
                 // ---------------------------------------------------
                 // GLOBAL
                 // If not local variable then check if global
                 // ---------------------------------------------------
                 // Variable definition should look like this:
                 // DEF GLOBAL DINT myVar_1 --> Create global integer var "myVar_1" 
                 //
                 // Token:
                 // [1] myVar_1
                 // [2]
                 // [3] DINT
                 // [4]
                 // [5] GLOBAL
                 // [6] 
                 // [7] DEF

                 // Init temp
                 #tempGlobal := FALSE;

                 // Check if number of token fits
                 IF #statTokenizedLine.numberOfToken = #statGlobalVariableDefinition.tokenizedString.numberOfToken THEN
                   // Set state initially --> Is overwritten in for loop
                   #statStateIntern := #STATE_LINE_IS_VAR_DEF;
                   #tempGlobal := TRUE;

                   // Check token of line to fit var declaration
                   FOR #tempCounter := 1 TO #statTokenizedLine.numberOfToken DO
                     // Skip name and type token
                     IF #tempCounter = #statGlobalVariableDefinition.nameTokenNumber
                       OR #tempCounter = #statGlobalVariableDefinition.typeTokenNumber
                     THEN
                       CONTINUE;
                       // Check the other keywords
                     ELSIF #statTokenizedLine.lineToken[#tempCounter] <> #statGlobalVariableDefinition.tokenizedString.lineToken[#tempCounter] THEN
                       // Mismatch between defintion and line 
                       // --> Not a variable definition
                       #statStateIntern := #STATE_IS_LINE_LABEL;
                       #tempGlobal := FALSE;
                       EXIT;
                     END_IF;
                   END_FOR;
                 ELSE
                   // Number of token does not fit
                   // Parse normal line
                   // Next step 
                   #statStateIntern := #STATE_IS_LINE_LABEL;
                   #tempGlobal := FALSE;
                 END_IF;

                 // Only check for local if not global
                 IF #tempGlobal = FALSE THEN
                   // ---------------------------------------------------
                   // LOCAL
                   // ---------------------------------------------------
                   // Variable definition should look like this:
                   // DEF DINT myVar_1 --> Create local integer var "myVar_1" 
                   //
                   // Token:
                   // [1] myVar_1
                   // [2]
                   // [3] DINT
                   // [4]
                   // [5] DEF

                   // Check if number of token fits
                   IF #statTokenizedLine.numberOfToken = #statLocalVariableDefinition.tokenizedString.numberOfToken THEN
                     // Set state initially --> Is overwritten in for loop
                     #statStateIntern := #STATE_LINE_IS_VAR_DEF;

                     // Check token of line to fit var declaration
                     FOR #tempCounter := 1 TO #statTokenizedLine.numberOfToken DO
                       // Skip name and type token
                       IF #tempCounter = #statLocalVariableDefinition.nameTokenNumber
                         OR #tempCounter = #statLocalVariableDefinition.typeTokenNumber
                       THEN
                         CONTINUE;
                         // Check the other keywords
                       ELSIF #statTokenizedLine.lineToken[#tempCounter] <> #statLocalVariableDefinition.tokenizedString.lineToken[#tempCounter] THEN
                         // Mismatch between defintion and line 
                         // --> Not a variable definition
                         #statStateIntern := #STATE_IS_LINE_LABEL;
                         EXIT;
                       END_IF;
                     END_FOR;
                   ELSE
                     // Number of token does not fit
                     // Parse normal line
                     // Next step 
                     #statStateIntern := #STATE_IS_LINE_LABEL;
                   END_IF;
                 END_IF;

               END_IF;

             END_REGION IS_LINE_VARIABLE_DEFINITION


             // ------------------------------------------------------------------------------------------
             // Line is variable definition
             // Line contains a variable definition like "DEF DINT myVar_1"
             // Go to STATE_LINE_PARSED
             // ------------------------------------------------------------------------------------------ 
             REGION LINE_IS_VARIABLE_DEFINITION
               IF #statStateIntern = #STATE_LINE_IS_VAR_DEF
               THEN
                 // Variable definition should look like this:
                 // DEF DINT myVar_1 --> Create local integer var "myVar_1" 
                 // Token:
                 // [1] myVar_1
                 // [2]
                 // [3] DINT
                 // [4]
                 // [5] DEF

                 // Check name to not be a number only!
                 IF NOT "LKinLang_IsTokenNumberInclSign"(#statTokenizedLine.lineToken[#statLocalVariableDefinition.nameTokenNumber]) THEN

                   // Check if name already exists as LABEL!
                   FOR #tempVarIndex := 1 TO #statLabelList.numberOfLabels DO
                     IF #statLabelList.labels[#tempVarIndex].labelName = #statTokenizedLine.lineToken[#statLocalVariableDefinition.nameTokenNumber] THEN
                       // Error: Variable already exists as label
                       #statStatus := #ERR_PARSING;
                       #statStateIntern := #STATE_ERROR;
                       #statErrorString := CONCAT(IN1 := #statErrorString, IN2 := 'Error: Variable already exists as label');
                       #statErrorString := CONCAT(IN1 := #statErrorString, IN2 := '; Line: ');
                       #statErrorString := CONCAT(IN1 := #statErrorString, IN2 := UDINT_TO_STRING(#statTokenizedLine.lineNo));
                       EXIT;
                     END_IF;
                   END_FOR;

                   // Check if name is a keyword
                   IF "LKinLang_IsTokenKeyWord"(token := #statTokenizedLine.lineToken[#statLocalVariableDefinition.nameTokenNumber], keyToken := #statKeyToken) THEN
                     // Error: Variable name can not be a keyword
                     #statStatus := #ERR_PARSING;
                     #statStateIntern := #STATE_ERROR;
                     #statErrorString := CONCAT(IN1 := #statErrorString, IN2 := 'Error: Variable name must not be a keyword');
                     #statErrorString := CONCAT(IN1 := #statErrorString, IN2 := '; Line: ');
                     #statErrorString := CONCAT(IN1 := #statErrorString, IN2 := UDINT_TO_STRING(#statTokenizedLine.lineNo));
                     EXIT;
                   END_IF;

                   // Check if name is a parameter 
                   FOR #tempVarIndex := 1 TO "LKINLANG_MAX_NUMBER_OF_PARAMETERS" DO
                     IF #statParameterLookUpTable[#tempVarIndex].parameterNameString = #statTokenizedLine.lineToken[#statLocalVariableDefinition.nameTokenNumber] THEN
                       // Error: Variable name can not be a keyword
                       #statStatus := #ERR_PARSING;
                       #statStateIntern := #STATE_ERROR;
                       #statErrorString := CONCAT(IN1 := #statErrorString, IN2 := 'Error: Variable name must not be a keyword');
                       #statErrorString := CONCAT(IN1 := #statErrorString, IN2 := '; Line: ');
                       #statErrorString := CONCAT(IN1 := #statErrorString, IN2 := UDINT_TO_STRING(#statTokenizedLine.lineNo));
                       EXIT;
                     END_IF;
                   END_FOR;

                   // Check if error occurred before
                   IF #statStateIntern <> #STATE_ERROR THEN
                     // Create local variable
                     // Imcrement local var counter
                     #statVarRefList.numberOfReferences += 1;

                     IF #statVarRefList.numberOfReferences > "LKINLANG_NUMBER_OF_VAR_REFS" THEN
                       // Error: Max number of variable references reached
                       #statStatus := #ERR_PARSING;
                       #statStateIntern := #STATE_ERROR;
                       #statErrorString := CONCAT(IN1 := #statErrorString, IN2 := 'Error: Overflow VarRefList; Increase NUMBER_OF_VAR_REFS');
                       #statErrorString := CONCAT(IN1 := #statErrorString, IN2 := '; Line: ');
                       #statErrorString := CONCAT(IN1 := #statErrorString, IN2 := UDINT_TO_STRING(#statTokenizedLine.lineNo));
                       EXIT;
                     ELSE
                       // Set step here because changing to error state could happen afterwards
                       // Next step --> Line finished
                       #statStateIntern := #STATE_LINE_PARSED;

                       // Copy name to table
                       #statVarRefList.references[#statVarRefList.numberOfReferences].name := #statTokenizedLine.lineToken[#statLocalVariableDefinition.nameTokenNumber];

                       // Check and set scope 
                       // Preset the scope to main
                       IF #tempGlobal = TRUE THEN
                         #statVarRefList.references[#statVarRefList.numberOfReferences].scope := 2; // Global var in main prg
                       ELSE
                         #statVarRefList.references[#statVarRefList.numberOfReferences].scope := 1; // Local var in main prg
                       END_IF;

                       // Iterate over subProgramList and check where we are currently
                       FOR #tempCounter := 1 TO #statSubPrgList.numberOfSubPrgs DO
                         IF #statTokenizedLine.lineNo > #statSubPrgList.subPrgs[#tempCounter].lineNumberStart
                           AND #statTokenizedLine.lineNo < #statSubPrgList.subPrgs[#tempCounter].lineNumberEnd
                         THEN
                           #statVarRefList.references[#statVarRefList.numberOfReferences].scope := #tempCounter * 10; // Local var in sub prg 
                           EXIT;
                         ELSIF #statTokenizedLine.lineNo < #statSubPrgList.subPrgs[#tempCounter].lineNumberStart THEN // Check if the current line number is smaller than the start of a sub --> Exit earlier
                           EXIT;
                         ELSE
                           CONTINUE;
                         END_IF;
                       END_FOR;

                       // Check if Global is allowed 
                       IF #tempGlobal = TRUE
                         AND #statVarRefList.references[#statVarRefList.numberOfReferences].scope >= 10
                       THEN
                         // Error: Not allowed to declare global in sub
                         #statStatus := #ERR_PARSING;
                         #statStateIntern := #STATE_ERROR;
                         #statErrorString := CONCAT(IN1 := #statErrorString, IN2 := 'Error: Declaring global variable in subprogram not allowed');
                         #statErrorString := CONCAT(IN1 := #statErrorString, IN2 := '; Line: ');
                         #statErrorString := CONCAT(IN1 := #statErrorString, IN2 := UDINT_TO_STRING(#statTokenizedLine.lineNo));
                         EXIT;
                       END_IF;

                       // Check if name already exists!
                       FOR #tempVarIndex := 1 TO #statVarRefList.numberOfReferences - 1 DO // exclude current entry
                         IF #statVarRefList.references[#tempVarIndex].name = #statVarRefList.references[#statVarRefList.numberOfReferences].name
                           AND #statVarRefList.references[#tempVarIndex].scope = #statVarRefList.references[#statVarRefList.numberOfReferences].scope
                         THEN
                           // Error: Variable already exists
                           #statStatus := #ERR_PARSING;
                           #statStateIntern := #STATE_ERROR;
                           #statErrorString := CONCAT(IN1 := #statErrorString, IN2 := 'Error: Variable already exists');
                           #statErrorString := CONCAT(IN1 := #statErrorString, IN2 := '; Line: ');
                           #statErrorString := CONCAT(IN1 := #statErrorString, IN2 := UDINT_TO_STRING(#statTokenizedLine.lineNo));
                           EXIT;
                         END_IF;
                       END_FOR;

                       // Decide type of variable
                       IF #statTokenizedLine.lineToken[#statLocalVariableDefinition.typeTokenNumber] = #statKeyToken.tokenBool THEN
                         #statVarRefList.references[#statVarRefList.numberOfReferences].type := "LKINLANG_VAR_TYPE_LOCAL_BOOL";
                         #statVariables.boolCounter += 1;
                         IF #statVariables.boolCounter > "LKINLANG_NUMBER_OF_LOCAL_BOOL" THEN
                           // Error too many local boolean
                           #statStatus := #ERR_PARSING;
                           #statStateIntern := #STATE_ERROR;
                           #statErrorString := CONCAT(IN1 := #statErrorString, IN2 := 'Error: Overflow local Bool; Increase "LKINLANG_NUMBER_OF_LOCAL_BOOL"');
                           #statErrorString := CONCAT(IN1 := #statErrorString, IN2 := '; Line: ');
                           #statErrorString := CONCAT(IN1 := #statErrorString, IN2 := UDINT_TO_STRING(#statTokenizedLine.lineNo));
                           EXIT;
                         ELSE
                           #statVarRefList.references[#statVarRefList.numberOfReferences].index := #statVariables.boolCounter;
                           #statVariables.boolean[#statVariables.boolCounter] := FALSE;
                         END_IF;
                       ELSIF #statTokenizedLine.lineToken[#statLocalVariableDefinition.typeTokenNumber] = #statKeyToken.tokenDInt THEN
                         #statVarRefList.references[#statVarRefList.numberOfReferences].type := "LKINLANG_VAR_TYPE_LOCAL_DINT";
                         #statVariables.dintCounter += 1;
                         IF #statVariables.dintCounter > "LKINLANG_NUMBER_OF_LOCAL_DINT" THEN
                           // Error too many local DInt
                           #statStatus := #ERR_PARSING;
                           #statStateIntern := #STATE_ERROR;
                           #statErrorString := CONCAT(IN1 := #statErrorString, IN2 := 'Error: Overflow local DInt; Increase "LKINLANG_NUMBER_OF_LOCAL_DINT"');
                           #statErrorString := CONCAT(IN1 := #statErrorString, IN2 := '; Line: ');
                           #statErrorString := CONCAT(IN1 := #statErrorString, IN2 := UDINT_TO_STRING(#statTokenizedLine.lineNo));
                           EXIT;
                         ELSE
                           #statVarRefList.references[#statVarRefList.numberOfReferences].index := #statVariables.dintCounter;
                           #statVariables.dints[#statVariables.dintCounter] := 0;
                         END_IF;
                       ELSIF #statTokenizedLine.lineToken[#statLocalVariableDefinition.typeTokenNumber] = #statKeyToken.tokenLReal THEN
                         #statVarRefList.references[#statVarRefList.numberOfReferences].type := "LKINLANG_VAR_TYPE_LOCAL_LREAL";
                         #statVariables.lrealCounter += 1;
                         IF #statVariables.lrealCounter > "LKINLANG_NUMBER_OF_LOCAL_LREAL" THEN
                           // Error too many local LReal
                           #statStatus := #ERR_PARSING;
                           #statStateIntern := #STATE_ERROR;
                           #statErrorString := CONCAT(IN1 := #statErrorString, IN2 := 'Error: Overflow local LReal; Increase "LKINLANG_NUMBER_OF_LOCAL_LREAL"');
                           #statErrorString := CONCAT(IN1 := #statErrorString, IN2 := '; Line: ');
                           #statErrorString := CONCAT(IN1 := #statErrorString, IN2 := UDINT_TO_STRING(#statTokenizedLine.lineNo));
                           EXIT;
                         ELSE
                           #statVarRefList.references[#statVarRefList.numberOfReferences].index := #statVariables.lrealCounter;
                           #statVariables.lreals[#statVariables.lrealCounter] := 0.0;
                         END_IF;
                       ELSE // type not defined
                         // Error wrong variable definition
                         #statStatus := #ERR_PARSING;
                         #statStateIntern := #STATE_ERROR;
                         #statErrorString := CONCAT(IN1 := #statErrorString, IN2 := 'Error: Type of local variable not defined');
                         #statErrorString := CONCAT(IN1 := #statErrorString, IN2 := '; Line: ');
                         #statErrorString := CONCAT(IN1 := #statErrorString, IN2 := UDINT_TO_STRING(#statTokenizedLine.lineNo));
                         EXIT;
                       END_IF;
                     END_IF;
                   ELSE
                     ;
                     // Error was already set
                     // --> do nothing
                   END_IF;

                 ELSE
                   // Error wrong variable definition
                   #statStatus := #ERR_PARSING;
                   #statStateIntern := #STATE_ERROR;
                   #statErrorString := CONCAT(IN1 := #statErrorString, IN2 := 'Error: Variable name can not be a number');
                   #statErrorString := CONCAT(IN1 := #statErrorString, IN2 := '; Line: ');
                   #statErrorString := CONCAT(IN1 := #statErrorString, IN2 := UDINT_TO_STRING(#statTokenizedLine.lineNo));
                   EXIT;
                 END_IF;
               END_IF;
             END_REGION LINE_IS_VARIABLE_DEFINITION

             // ------------------------------------------------------------------------------------------
             // Is line label
             // Check if the line contains a correct LABEL
             // YES: Go to STATE_LINE_PARSED
             // NO: Go to IS_LINE_GOTO 
             // ------------------------------------------------------------------------------------------ 
             REGION IS_LINE_LABEL
               IF #statStateIntern = #STATE_IS_LINE_LABEL
               THEN
                 // Check if line starts with 'LABEL'
                 IF #statTokenizedLine.lineToken[#statTokenizedLine.numberOfToken] = #statKeyToken.tokenJumpTarget THEN

                   // Nothing to do when token is LABEL as the labelList was already created
                   #statStateIntern := #STATE_LINE_PARSED;

                   // Create LabelList at runtime here
                   (*
                   // Check if line contains exactly 3 tokens
                   // Definition:
                   // [1] "myLabel"
                   // [2] " "
                   // [3] "LABEL"
                   IF #statTokenizedLine.numberOfToken = 3
                     AND #statTokenizedLine.LineToken[#statTokenizedLine.numberOfToken - 1] = ' ' // second token must be space
                     AND NOT "LKinLang_IsTokenNumber"(#statTokenizedLine.LineToken[#statTokenizedLine.numberOfToken - 2]) // first token must not be a number
                   THEN
                     ; // correct label definition 
                     // Reset bit
                     #tempLabelExists := FALSE;
                     // Check labelList if label already exists
                     FOR #tempCounter := 1 TO #statLabelList.numberOfLabels DO
                       IF #statLabelList.labels[#tempCounter].labelName = #statTokenizedLine.LineToken[#statTokenizedLine.numberOfToken - 2]
                       THEN
                         //Check if the line numbers are different 
                         IF #statLabelList.labels[#tempCounter].lineNumber <> #statTokenizedLine.lineNo 
                         THEN
                           // Label already exists in other line
                           // Throw error
                           #statStatus := #ERR_PARSING;
                           #statStateIntern := #STATE_ERROR;
                           #statErrorString := CONCAT(IN1 := #statErrorString, IN2 := ';Error: Label is not unique');
                           #statErrorString := CONCAT(IN1 := #statErrorString, IN2 := ' in line: ');
                           #statErrorString := CONCAT(IN1 := #statErrorString, IN2 := UDINT_TO_STRING(#statTokenizedLine.lineNo));
                           EXIT;
                         ELSE
                           // Label is already in list 
                           // But with same line number 
                           // Maybe jumped back and found same label again
                           // --> No error just dont add again
                           // Set bit to signal label already exists
                           #tempLabelExists := TRUE;
                           // Go to LineParsed
                           #statStateIntern := #STATE_LINE_PARSED;
                           EXIT;
                         END_IF;
                       END_IF;
                     END_FOR;

                     // Check if the number of labels is ok 
                     IF #statLabelList.numberOfLabels >= "LKINLANG_NUMBER_OF_LABELS" AND #tempLabelExists = FALSE THEN
                       // No more space in labelList
                       // Throw error 
                       #statStatus := #ERR_PARSING;
                       #statStateIntern := #STATE_ERROR;
                       #statErrorString := CONCAT(IN1 := #statErrorString, IN2 := ';Error: Maximum number of labels reached');
                       #statErrorString := CONCAT(IN1 := #statErrorString, IN2 := ' in line: ');
                       #statErrorString := CONCAT(IN1 := #statErrorString, IN2 := UDINT_TO_STRING(#statTokenizedLine.lineNo));
                       EXIT;
                     END_IF;

                     IF #statStateIntern <> #STATE_ERROR AND #tempLabelExists = FALSE THEN
                       // Increment number of labels if possible
                       #statLabelList.numberOfLabels += 1;
                       // Set the label info
                       #statLabelList.labels[#statLabelList.numberOfLabels].labelName := #statTokenizedLine.LineToken[#statTokenizedLine.numberOfToken - 2];
                       #statLabelList.labels[#statLabelList.numberOfLabels].lineNumber := #statTokenizedLine.lineNo;
                       // TODO: Add hierarchic level?
                       // 
                       // Go to LineParsed
                       #statStateIntern := #STATE_LINE_PARSED;
                     ELSE
                       // Error was set already set
                       // Do nothing
                       ;
                     END_IF;


                   ELSE
                     // Wrong label definition 
                     // Throw error
                     #statStatus := #ERR_PARSING;
                     #statStateIntern := #STATE_ERROR;
                     #statErrorString := CONCAT(IN1 := #statErrorString, IN2 := ';Error: Invalid label definition');
                     #statErrorString := CONCAT(IN1 := #statErrorString, IN2 := ' in line: ');
                     #statErrorString := CONCAT(IN1 := #statErrorString, IN2 := UDINT_TO_STRING(#statTokenizedLine.lineNo));
                     EXIT;
                   END_IF;
                   *)


                 ELSE
                   // Not a label definition
                   // Go to next state
                   #statStateIntern := #STATE_IS_LINE_GOTO;
                 END_IF;
               END_IF;


             END_REGION IS_LINE_LABEL

             // ------------------------------------------------------------------------------------------
             // Is line GOTO, GOTOC
             // Check if the line contains a GOTO, GOTOC, ...
             // If yes then set the next lineNumber to be parsed
             // YES: Go to STATE_LINE_PARSED
             // NO: Go to IS_LINE_STOPRE
             // ------------------------------------------------------------------------------------------ 
             REGION IS_LINE_GOTO
               IF #statStateIntern = #STATE_IS_LINE_GOTO
               THEN
                 // Check if line starts with 'GOTO'
                 IF (#statTokenizedLine.lineToken[#statTokenizedLine.numberOfToken] = #statKeyToken.tokenJump AND #statTokenizedLine.numberOfToken = 3)
                   OR #statTokenizedLine.lineToken[#statTokenizedLine.numberOfToken] = #statKeyToken.tokenJumpConditional
                 THEN
                   // Definition GOTO:             // Definition GOTOC:
                   // [1] "myLabel"                // [1] "10"
                   // [2] " "                      // [2] ">"
                   // [3] "GOTO"                   // [3] "counter"
                   //                              // [4] " "
                   //                              // [5] "myLabel"
                   //                              // [6] " "
                   //                              // [7] "GOTOC"

                   IF #statTokenizedLine.lineToken[#statTokenizedLine.numberOfToken - 1] = ' ' // second token must be space
                     AND NOT "LKinLang_IsTokenNumberInclSign"(#statTokenizedLine.lineToken[#statTokenizedLine.numberOfToken - 2]) // labelName must not be a number
                   THEN
                     // correct jump definition 
                     // Check labelList if label exists
                     #tempLabelExists := FALSE;
                     FOR #tempLabelIndex := 1 TO #statLabelList.numberOfLabels DO
                       IF #statLabelList.labels[#tempLabelIndex].labelName = #statTokenizedLine.lineToken[#statTokenizedLine.numberOfToken - 2] THEN
                         // Label exists!
                         // Exit this loop
                         #tempLabelExists := TRUE;
                         EXIT;
                       END_IF;
                     END_FOR;

                     IF #tempLabelExists THEN
                       // Check if GOTO or GOTOC
                       // And get condition result
                       IF #statTokenizedLine.lineToken[#statTokenizedLine.numberOfToken] = #statKeyToken.tokenJump THEN
                         #tempConditionResult := TRUE;
                       ELSE
                         // correct jump definition 
                         // Evaluate condition 
                         // Evaluate the condition after the label name to decide if the jump is executed or not
                         // Evaluation could work like normal parse line tokens?
                         #tempConditionResult := "LKinLang_EvaluateCondition"(offsetLastTokenIndex := 3, // Token offset where condition begins
                                                                              tokenizedLine := #statTokenizedLine,
                                                                              varRefList := #statVarRefList,
                                                                              localVariables := #statVariables,
                                                                              interfaceVariables := #interfaceVariables,
                                                                              keyToken := #statKeyToken,
                                                                              subPrgList := #statSubPrgList,
                                                                              errorString := #statErrorString);


                         // Check if error occured in FC
                         IF #statErrorString <> '' THEN
                           #statStatus := #ERR_PARSING;
                           #statStateIntern := #STATE_ERROR;
                           // Error string was already set
                         END_IF;
                       END_IF;

                       // In case of syntaxCheck being on, always set the condition result to false 
                       // --> Avoid jumping 
                       IF #statSyntaxCheck <> "LKINLANG_SYNTAX_CHECK_OFF" THEN
                         #tempConditionResult := FALSE;
                       END_IF;

                       IF #tempConditionResult AND #statStateIntern <> #STATE_ERROR THEN
                         // Check if jump to label is allowed 
                         // Get current hierarchicLevel
                         #statHierarchicLevel.currentLevel := 0;
                         FOR #tempCounter := 1 TO #statHierarchicLevel.numberOfLevels DO
                           IF #statTokenizedLine.lineNo >= #statHierarchicLevel.levels[#tempCounter].lineNumber THEN
                             #statHierarchicLevel.currentLevel := #statHierarchicLevel.levels[#tempCounter].level;
                           ELSE
                             EXIT;
                           END_IF;
                         END_FOR;

                         // Check if jumping from main to sub
                         IF #statTokenizedLine.lineNo < #statSubPrgList.subPrgs[1].lineNumberStart
                           AND #statLabelList.labels[#tempLabelIndex].lineNumber >= #statSubPrgList.subPrgs[1].lineNumberStart
                         THEN
                           // Throw error --> Not allowed to jump between programs
                           #statStatus := #ERR_PARSING;
                           #statStateIntern := #STATE_ERROR;
                           #statErrorString := CONCAT(IN1 := #statErrorString, IN2 := 'Error: Jump from main to subprogram not allowed');
                           #statErrorString := CONCAT(IN1 := #statErrorString, IN2 := ' in line: ');
                           #statErrorString := CONCAT(IN1 := #statErrorString, IN2 := UDINT_TO_STRING(#statTokenizedLine.lineNo));
                           EXIT;
                         END_IF;


                         // Check if current level is greater or equal else throw error! 
                         // Jumps are only allowed if target is not in a different loop?
                         IF #statHierarchicLevel.currentLevel >= #statLabelList.labels[#tempLabelIndex].hierarchicLevel THEN
                           // Remove stack entry which are left
                           FOR #tempCounter := #statStack.numberOfElements TO 1 BY -1 DO
                             // Check if Label is outside of subprogram --> Throw error --> Not allowed
                             IF #statStack.stackElements[#tempCounter].type = "LKINLANG_ENTRY_TYPE_SUB" THEN
                               IF #statLabelList.labels[#tempLabelIndex].lineNumber < #statSubPrgList.subPrgs[#statStack.stackElements[#tempCounter].quantity].lineNumberStart
                                 OR #statLabelList.labels[#tempLabelIndex].lineNumber > #statSubPrgList.subPrgs[#statStack.stackElements[#tempCounter].quantity].lineNumberEnd
                               THEN
                                 // Throw error --> Not allowed to jump between programs
                                 #statStatus := #ERR_PARSING;
                                 #statStateIntern := #STATE_ERROR;
                                 #statErrorString := CONCAT(IN1 := #statErrorString, IN2 := 'Error: Jump between programs not allowed');
                                 #statErrorString := CONCAT(IN1 := #statErrorString, IN2 := ' in line: ');
                                 #statErrorString := CONCAT(IN1 := #statErrorString, IN2 := UDINT_TO_STRING(#statTokenizedLine.lineNo));
                                 EXIT;
                               END_IF;
                             END_IF;

                             // Check if the target line number is before or after a stack entry --> Leaving loop --> Delete stack entry
                             IF #statLabelList.labels[#tempLabelIndex].lineNumber > #statStack.stackElements[#tempCounter].lineNumberEnd
                               OR #statLabelList.labels[#tempLabelIndex].lineNumber < #statStack.stackElements[#tempCounter].lineNumberStart
                             THEN
                               // Delete stack entry
                               #statStack.stackElements[#tempCounter].lineNumberStart := 0;
                               #statStack.stackElements[#tempCounter].lineNumberEnd := 0;
                               #statStack.stackElements[#tempCounter].type := 0;
                               #statStack.stackElements[#tempCounter].increment := 0;
                               #statStack.stackElements[#tempCounter].quantity := 0;
                               #statStack.stackElements[#tempCounter].variableRef.index := 0;
                               #statStack.stackElements[#tempCounter].variableRef.type := 0;
                               #statStack.stackElements[#tempCounter].variableRef.name := '';
                               // Count one backwards
                               #statStack.numberOfElements -= 1;
                             END_IF;
                           END_FOR;

                           // Only request line if no error occured
                           IF #statStateIntern <> #STATE_ERROR THEN
                             // Go to line containing LABEL 
                             #statSearchedLine := #statLabelList.labels[#tempLabelIndex].lineNumber;
                             #statStateIntern := #STATE_LINE_PARSED;
                           END_IF;
                         ELSE
                           // ERROR jump not allowed
                           #statStatus := #ERR_PARSING;
                           #statStateIntern := #STATE_ERROR;
                           #statErrorString := CONCAT(IN1 := #statErrorString, IN2 := 'Error: Jump to lower level is not allowed');
                           #statErrorString := CONCAT(IN1 := #statErrorString, IN2 := ' in line: ');
                           #statErrorString := CONCAT(IN1 := #statErrorString, IN2 := UDINT_TO_STRING(#statTokenizedLine.lineNo));
                           EXIT;
                         END_IF;

                       ELSE
                         // Condition is false 
                         // --> No jump!
                         // Line finished
                         #statStateIntern := #STATE_LINE_PARSED;
                       END_IF;
                     ELSE
                       // Error label does not exist
                       // Throw error
                       #statStatus := #ERR_PARSING;
                       #statStateIntern := #STATE_ERROR;
                       #statErrorString := CONCAT(IN1 := #statErrorString, IN2 := ';Error: Jump target does not exist');
                       #statErrorString := CONCAT(IN1 := #statErrorString, IN2 := ' in line: ');
                       #statErrorString := CONCAT(IN1 := #statErrorString, IN2 := UDINT_TO_STRING(#statTokenizedLine.lineNo));
                       EXIT;
                     END_IF;

                   ELSE
                     // Wrong jump definition 
                     // Throw error
                     #statStatus := #ERR_PARSING;
                     #statStateIntern := #STATE_ERROR;
                     #statErrorString := CONCAT(IN1 := #statErrorString, IN2 := ';Error: Invalid jump definition');
                     #statErrorString := CONCAT(IN1 := #statErrorString, IN2 := ' in line: ');
                     #statErrorString := CONCAT(IN1 := #statErrorString, IN2 := UDINT_TO_STRING(#statTokenizedLine.lineNo));
                     EXIT;
                   END_IF;
                 ELSE
                   // Not a jump definition
                   // Go to next state
                   #statStateIntern := #STATE_IS_LINE_STOPRE;
                 END_IF;
               END_IF;

             END_REGION IS_LINE_GOTO

             // ------------------------------------------------------------------------------------------
             // Is line STOPRE
             // Check if the line contains STOPRE
             // If yes then signalize to MovePath and wait with parsing
             // YES: Go to STATE_PREPROCESSING_STOP
             // NO: Go to IS_LINE_IF
             // ------------------------------------------------------------------------------------------ 
             REGION IS_LINE_STOPRE
               IF #statStateIntern = #STATE_IS_LINE_STOPRE
               THEN
                 // Check if line starts with 'STOPRE' and contains 1 token
                 IF #statTokenizedLine.lineToken[#statTokenizedLine.numberOfToken] = #statKeyToken.tokenPreprocessingStop
                   AND #statTokenizedLine.numberOfToken = 1
                 THEN
                   // Only set STOPRE if syntac check if off
                   IF #statSyntaxCheck = "LKINLANG_SYNTAX_CHECK_OFF" THEN
                     // Set stopre bit for movePath and switch state to interrupt parsing until movePath catches up
                     #pathData.pointers.preprocessingStop := TRUE;
                     // Unlock buffer if locked --> Stopre in first few commands
                     #pathData.pointers.bufferLocked := FALSE;
                     #statStateIntern := #STATE_PREPROCESSING_STOP;
                   ELSE
                     // Line is parsed
                     #statStateIntern := #STATE_LINE_PARSED;
                   END_IF;
                 ELSE
                   // Check if line contains IF
                   #statStateIntern := #STATE_IS_LINE_IF;
                 END_IF;
               END_IF;
             END_REGION IS_LINE_STOPRE

             // ------------------------------------------------------------------------------------------
             // Is line IF
             // Check if the line contains IF, ELSE or ENDIF
             // If yes then evaluate condtion and continue accordingly
             // YES: Go to STATE_LINE_PARSED
             // NO: Go to IS_LINE_WHILE
             // ------------------------------------------------------------------------------------------ 
             REGION IS_LINE_IF
               IF #statStateIntern = #STATE_IS_LINE_IF
               THEN
                 // Definition IF:
                 // [1] "10"
                 // [2] ">"
                 // [3] "counter"
                 // [4] " "
                 // [5] "IF"

                 // Check if line starts with 'IF'
                 IF #statTokenizedLine.lineToken[#statTokenizedLine.numberOfToken] = #statKeyToken.tokenIf THEN
                   REGION IF
                     // IF is found
                     #statStack.numberOfElements += 1;
                     IF #statStack.numberOfElements <= "LKINLANG_NUMBER_OF_STACK_ELEMENTS" THEN
                       #statStack.stackElements[#statStack.numberOfElements].type := "LKINLANG_ENTRY_TYPE_IF";
                       #statStack.stackElements[#statStack.numberOfElements].lineNumberStart := #statTokenizedLine.lineNo;
                     ELSE
                       // Error Stack overflow
                       #statStatus := #ERR_PARSING;
                       #statStateIntern := #STATE_ERROR;
                       #statErrorString := CONCAT(IN1 := #statErrorString, IN2 := 'Error: Maximum array index of stack reached');
                       #statErrorString := CONCAT(IN1 := #statErrorString, IN2 := ' in line: ');
                       #statErrorString := CONCAT(IN1 := #statErrorString, IN2 := UDINT_TO_STRING(#statTokenizedLine.lineNo));
                     END_IF;

                     IF #statStateIntern <> #STATE_ERROR THEN
                       // Evaluate the condition and decide where to go next
                       #tempConditionResult := "LKinLang_EvaluateCondition"(offsetLastTokenIndex := 2, // Token offset where condition begins
                                                                            tokenizedLine := #statTokenizedLine,
                                                                            varRefList := #statVarRefList,
                                                                            localVariables := #statVariables,
                                                                            interfaceVariables := #interfaceVariables,
                                                                            keyToken := #statKeyToken,
                                                                            subPrgList := #statSubPrgList,
                                                                            errorString := #statErrorString);


                       // Check if error occured in FC
                       IF #statErrorString <> '' THEN
                         #statStatus := #ERR_PARSING;
                         #statStateIntern := #STATE_ERROR;
                         // Error string was already set
                       END_IF;
                     END_IF;

                     // Check if error occured
                     IF #statStateIntern <> #STATE_ERROR THEN
                       // Check for ENDIF
                       // Search current level of IF and find matching EndIF  
                       #tempConditionCounter := -1;
                       FOR #tempCounter := 1 TO #statHierarchicLevel.numberOfLevels DO
                         IF #statHierarchicLevel.levels[#tempCounter].lineNumber = #statTokenizedLine.lineNo THEN
                           #tempConditionCounter := #statHierarchicLevel.levels[#tempCounter].level; // This is the hierarchic level of the current IF
                           CONTINUE;
                         END_IF;

                         IF #statHierarchicLevel.levels[#tempCounter].type = "LKINLANG_ENTRY_TYPE_ENDIF"
                           AND #statHierarchicLevel.levels[#tempCounter].level = #tempConditionCounter THEN
                           // Correct endIF found
                           // Exit for loop
                           #tempLineNumber := #statHierarchicLevel.levels[#tempCounter].lineNumber;
                           EXIT;
                         END_IF;
                       END_FOR;

                       // Check if token for ENDIF was found
                       IF #tempLineNumber <= 0 THEN
                         // Error no ENDIF found to IF
                         #statStatus := #ERR_PARSING;
                         #statStateIntern := #STATE_ERROR;
                         #statErrorString := CONCAT(IN1 := #statErrorString, IN2 := 'Error: No matching ');
                         #statErrorString := CONCAT(IN1 := #statErrorString, IN2 := #statKeyToken.tokenEndIf);
                         #statErrorString := CONCAT(IN1 := #statErrorString, IN2 := ' found to ');
                         #statErrorString := CONCAT(IN1 := #statErrorString, IN2 := #statKeyToken.tokenIf);
                         #statErrorString := CONCAT(IN1 := #statErrorString, IN2 := ' in line: ');
                         #statErrorString := CONCAT(IN1 := #statErrorString, IN2 := UDINT_TO_STRING(#statTokenizedLine.lineNo));
                       END_IF;

                       // Check if error was set
                       IF #statStateIntern <> #STATE_ERROR THEN

                         // In case of syntaxCheck being on, always set the condition result to true 
                         // --> Always check if condition
                         IF #statSyntaxCheck <> "LKINLANG_SYNTAX_CHECK_OFF" THEN
                           #tempConditionResult := TRUE;
                         END_IF;

                         // Check the result of the condition
                         IF #tempConditionResult = FALSE THEN
                           // Condition is false --> check for ELSE
                           // Search current level of IF and find matching ELSE
                           #tempConditionCounter := -1;
                           FOR #tempCounter := 1 TO #statHierarchicLevel.numberOfLevels DO
                             IF #statHierarchicLevel.levels[#tempCounter].lineNumber = #statTokenizedLine.lineNo THEN
                               #tempConditionCounter := #statHierarchicLevel.levels[#tempCounter].level; // This is the hierarchic level of the current IF
                               CONTINUE;
                             END_IF;

                             // Check if the lineNumber is already greater than the ENDIF we found
                             IF #statHierarchicLevel.levels[#tempCounter].lineNumber > #tempLineNumber THEN
                               // No matching else found
                               EXIT;
                             END_IF;

                             IF #statHierarchicLevel.levels[#tempCounter].type = "LKINLANG_ENTRY_TYPE_ELSE"
                               AND #statHierarchicLevel.levels[#tempCounter].level = #tempConditionCounter THEN
                               // Correct ELSE found
                               // Exit for loop
                               #tempLineNumber := #statHierarchicLevel.levels[#tempCounter].lineNumber + 1;
                               EXIT;
                             END_IF;
                           END_FOR;

                           // Go to line after ELSE or line containing ENDIF
                           #statSearchedLine := #tempLineNumber;
                           #statStateIntern := #STATE_LINE_PARSED;
                         ELSE
                           // Condition is TRUE and ENDIF is ok --> Nothing more to do
                           #statStateIntern := #STATE_LINE_PARSED;
                         END_IF;
                       END_IF;
                     END_IF;
                   END_REGION IF

                 ELSIF #statTokenizedLine.lineToken[#statTokenizedLine.numberOfToken] = #statKeyToken.tokenElse
                   AND #statTokenizedLine.numberOfToken = 1
                 THEN
                   REGION ELSE
                     // Else found
                     // If we reach this condition then the previous IF condition was true --> Skip this else part and search endIf
                     // Check if the previos stack entry was a IF and if there are elements on the stack
                     IF #statStack.numberOfElements > 0 THEN
                       IF #statStack.stackElements[#statStack.numberOfElements].type = "LKINLANG_ENTRY_TYPE_IF" THEN
                         // Search current level of IF and find matching ENDIF  
                         #tempConditionCounter := -1;
                         FOR #tempCounter := 1 TO #statHierarchicLevel.numberOfLevels DO
                           IF #statHierarchicLevel.levels[#tempCounter].lineNumber = #statTokenizedLine.lineNo THEN
                             #tempConditionCounter := #statHierarchicLevel.levels[#tempCounter].level; // This is the hierarchic level of the current IF
                             CONTINUE;
                           END_IF;

                           IF #statHierarchicLevel.levels[#tempCounter].type = "LKINLANG_ENTRY_TYPE_ENDIF"
                             AND #statHierarchicLevel.levels[#tempCounter].level = #tempConditionCounter THEN
                             // Correct ENDIF found
                             #tempLineNumber := #statHierarchicLevel.levels[#tempCounter].lineNumber;
                             EXIT;
                           END_IF;
                         END_FOR;

                         // If syntax check is not off then continue in next line
                         IF #statSyntaxCheck = "LKINLANG_SYNTAX_CHECK_OFF" THEN
                           // Goto line containing "ENDIF" 
                           #statSearchedLine := #tempLineNumber;
                           #statStateIntern := #STATE_LINE_PARSED;
                         ELSE
                           // Go to next state
                           #statStateIntern := #STATE_LINE_PARSED;
                         END_IF;

                       ELSE
                         // Error last entry on stack was not an IF
                         #statStatus := #ERR_PARSING;
                         #statStateIntern := #STATE_ERROR;
                         #statErrorString := CONCAT(IN1 := #statErrorString, IN2 := 'Error: No matching ');
                         #statErrorString := CONCAT(IN1 := #statErrorString, IN2 := #statKeyToken.tokenIf);
                         #statErrorString := CONCAT(IN1 := #statErrorString, IN2 := ' found to ');
                         #statErrorString := CONCAT(IN1 := #statErrorString, IN2 := #statKeyToken.tokenElse);
                         #statErrorString := CONCAT(IN1 := #statErrorString, IN2 := ' in line: ');
                         #statErrorString := CONCAT(IN1 := #statErrorString, IN2 := UDINT_TO_STRING(#statTokenizedLine.lineNo));
                       END_IF;
                     ELSE
                       // Error no more elements on stack
                       #statStatus := #ERR_PARSING;
                       #statStateIntern := #STATE_ERROR;
                       #statErrorString := CONCAT(IN1 := #statErrorString, IN2 := 'Error: ');
                       #statErrorString := CONCAT(IN1 := #statErrorString, IN2 := #statKeyToken.tokenElse);
                       #statErrorString := CONCAT(IN1 := #statErrorString, IN2 := ' not allowed in line: ');
                       #statErrorString := CONCAT(IN1 := #statErrorString, IN2 := UDINT_TO_STRING(#statTokenizedLine.lineNo));
                     END_IF;
                   END_REGION ELSE

